// Mitsubishi GX Works2 project: Calculate   PLC: Q06UDEH (continued)

Import2Switch(ConveyorEntryIO:=Import2SwitchConveyorIn,
                          ConveyorExitIO:=Import2SwitchConveyorOut ,
                           SwitchIO:=Import2SwitchIO);
Import2SwitchIO.xLiftCylinderExtendButton:=M155;
Import2SwitchIO.xLiftCylinderRetractButton:=M156;
Y1ED:=Import2SwitchIO.xLiftCylinderExtend;
Y1EE:=Import2SwitchIO.xLiftCylinderRetract;
Import2SwitchIO.xLiftCylinderExtendDetect:=XF1;
Import2SwitchIO.xLiftCylinderRetractDetect:=XF2;
Import2SwitchConveyorIn.xCWPresent:=X104;
Import2SwitchConveyorIn.tLoadDelay:=T#2s;
Import2SwitchConveyorOut.xForward:=M149;
Import2SwitchConveyorOut.tLeaveDelay:=t#8s;
Import2SwitchConveyorOut.xCWPresent:=XF0;
Y1FC:=Import2SwitchConveyorIn.xMotorCW;

Import2LoadCylinder(ShuttleCarInOut:=Import2LoadCylinderIO);
ShuttleCarCurrentPosition( XF6 OR XF7 ,XF6 ,XF7, FALSE, Import2LoadCylinderIO.iCurrentPos );
Import2LoadCylinderIO.xReady:=TRUE;
Import2LoadCylinderIO.xForward:=M161;
Import2LoadCylinderIO.xBackward:=M162;
Import2LoadCylinderIO.xPosLimit:=TRUE;
Import2LoadCylinderIO.xNegLimit:=TRUE;
Y1ED:=Import2LoadCylinderIO.xCW;
Y1EE:=Import2LoadCylinderIO.xCCW;

(*2巷道出库*)
Export2Conveyor1(ConveyorMotor:=Export2Conveyor1IO);
Export2Conveyor1IO.tLeaveDelay:=t#10s;
Export2Conveyor1IO.xForward:=M96;
Export2Conveyor1IO.xCWPresent:=XFB;
Y1FD:=Export2Conveyor1IO.xMotorCW;

Export2Conveyor2(ConveyorMotor:=Export2Conveyor2iO);
Export2Conveyor2IO.tLeaveDelay:=t#10s;
Export2Conveyor2IO.xForward:=M97;
Export2Conveyor2IO.xCWPresent:=XFC;
Y1FE:=Export2Conveyor2IO.xMotorCW;

Export2Switch(ConveyorEntryIO:=Export2SwitchConveyorIn,
                          ConveyorExitIO:=Export2SwitchConveyorOut ,
                           SwitchIO:=Export2SwitchIO);
Export2SwitchIO.xLiftCylinderExtendButton:=M120;
Export2SwitchIO.xLiftCylinderRetractButton:=M121;
Export2SwitchIO.xLiftCylinderExtendInit:=1;
Y1F1:=Export2SwitchIO.xLiftCylinderExtend;
Y1F0:=Export2SwitchIO.xLiftCylinderRetract;
Export2SwitchIO.xLiftCylinderExtendDetect:=XF9;
Export2SwitchIO.xLiftCylinderRetractDetect:=XFA;
Export2SwitchConveyorIn.xForward:=M123;
Export2SwitchConveyorIn.xCWPresent:=X105;
Y1FF:=Export2SwitchConveyorIn.xMotorCW;
Export2SwitchConveyorOut.xCWPresent:=X105;

Export2LoadCylinder(ShuttleCarInOut:=Export2LoadCylinderIO);
ShuttleCarCurrentPosition( XFF OR XFE ,XFF ,XFE, FALSE, Export2LoadCylinderIO.iCurrentPos );
Export2LoadCylinderIO.xReady:=TRUE;
Export2LoadCylinderIO.xForward:=M124;
Export2LoadCylinderIO.xBackward:=M125;
Export2LoadCylinderIO.xPosLimit:=TRUE;
Export2LoadCylinderIO.xNegLimit:=TRUE;
Y1F2:=Export2LoadCylinderIO.xCW;
Y1F3:=Export2LoadCylinderIO.xCCW;

IF g_xAuto THEN
	(**高温库前自动程序**)
	Y187:=1;(***出库倍速链***)
(*	Y186:=1;(***入库倍速链***)
	IF  M883 AND XED THEN
        Export1LoadCylinderIO.xMDIExe:=1;
        Export1LoadCylinderIO.iDestinationPos:=1;
	END_IF;
	IF NOT XED THEN
        Export1LoadCylinderIO.xMDIExe:=1;
        Export1LoadCylinderIO.iDestinationPos:=2;
     END_IF;		
	Export1Conveyor1IO.xLoad:=XED AND Export1LoadCylinderIO.iCurrentPos=2;
	Export1Conveyor1IO.xUnload:=Export1Conveyor2IO.xEmpty;
	Export1Conveyor2IO.xLoad:=Export1Conveyor1IO.xNextRun;
	IF Y1E5 THEN
		Export1SwitchIO.xLiftCylinderExtendInit:=0;
	ELSE
		Export1SwitchIO.xLiftCylinderExtendInit:=1;
	END_IF;
	Export1Conveyor2Io.xUnload:=Export1SwitchConveyorIn.xEmpty;
	Export1SwitchIO.xEntryEnable:=Export1Conveyor2Io.xNextRun;
	Export1SwitchIO.xSwithEnable:=1;
	IF  M884 THEN
        Export2LoadCylinderIO.xMDIExe:=1;
        Export2LoadCylinderIO.iDestinationPos:=2;
	END_IF;
	Export2Conveyor1IO.xLoad:=XFD AND Export2LoadCylinderIO.iCurrentPos=2;
	Export2Conveyor1IO.xUnload:=Export2Conveyor2IO.xEmpty;
	Export2Conveyor2IO.xLoad:=Export2Conveyor1IO.xNextRun;
	Export2Conveyor2Io.xUnload:=Export2SwitchConveyorIn.xEmpty;
	Export2SwitchIO.xEntryEnable:=Export2Conveyor2Io.xNextRun;
	Export2SwitchIO.xSwithEnable:=1;
	
	H3000SwitchQuadPackageIO.xEntryEnable:=1;
	H3000SwitchQuadPackageIO.xSwithEnable:=1;
	H3000SwitchQuadPackageio.xExitEnable:=H3000Conveyor1IO.xEmpty;
	H3000Conveyor1Io.xLoad:=H3000SwitchPackageConveyorOut.xNextRun;
	H3000Conveyor1IO.xUnload:=H3000Conveyor2IO.xEmpty;
	H3000Conveyor2IO.xLoad:=H3000Conveyor1IO.xNextRun;
	H3000Conveyor2IO.xUnload:=H3000Conveyor3IO.xEmpty;
	H3000Conveyor3IO.xLoad:=H3000Conveyor2IO.xNextRun;	
	H3000Conveyor3IO.xUnload:=H3000Conveyor4IO.xEmpty;
	H3000Conveyor4IO.xLoad:=H3000Conveyor3IO.xNextRun;
	H3000Conveyor4IO.xUnload:=H3000Conveyor5IO.xEmpty;
	H3000Conveyor5IO.xLoad:=H3000Conveyor4IO.xNextRun;
	H3000Conveyor5IO.xUnload:=H3000Conveyor6IO.xEmpty;
	H3000Conveyor6IO.xLoad:=H3000Conveyor5IO.xNextRun;
	H3000Conveyor6IO.xUnload:=H3000Conveyor7IO.xEmpty;
	H3000Conveyor7IO.xLoad:=H3000Conveyor6IO.xNextRun;
	H3000Conveyor7IO.xUnload:=H3000Conveyor8IO.xEmpty;
	H3000Conveyor8IO.xLoad:=H3000Conveyor7IO.xNextRun;	
	H3000Conveyor8IO.xUnload:=H3000Conveyor9IO.xEmpty;
	H3000Conveyor9IO.xLoad:=H3000Conveyor8IO.xNextRun;	
	H3000Conveyor9IO.xUnload:=H3000Conveyor10IO.xEmpty;
	H3000Conveyor10IO.xLoad:=H3000Conveyor9IO.xNextRun;
	H3000Conveyor10IO.xUnload:=D401.0;
	D201.0:=H3000Conveyor10IO.xNextRun;

	
	(*H2200Conveyor1IO.xLoad:=;*)
	H2200Conveyor1IO.xUnload:=H2200Conveyor2IO.xEmpty;
	H2200Conveyor2IO.xLoad:=H2200Conveyor1IO.xNextRun;
	H2200Conveyor2IO.xUnload:=H2200Conveyor3IO.xEmpty;
	H2200Conveyor3IO.xLoad:=H2200Conveyor2IO.xNextRun;	
	H2200Conveyor3IO.xUnload:=H2200Conveyor4IO.xEmpty;
	H2200Conveyor4IO.xLoad:=H2200Conveyor3IO.xNextRun;
	H2200Conveyor4IO.xUnload:=H2200Conveyor5IO.xEmpty;
	H2200Conveyor5IO.xLoad:=H2200Conveyor4IO.xNextRun;
	H2200Conveyor5IO.xUnload:=H2200Conveyor6IO.xEmpty;
	H2200Conveyor6IO.xLoad:=H2200Conveyor5IO.xNextRun;
	H2200Conveyor6IO.xUnload:=H2200Conveyor7IO.xEmpty;
	H2200Conveyor7IO.xLoad:=H2200Conveyor6IO.xNextRun;
	H2200Conveyor7IO.xUnload:=H2200Conveyor8IO.xEmpty;
	H2200Conveyor8IO.xLoad:=H2200Conveyor7IO.xNextRun;	
	H2200Conveyor8IO.xUnload:=H2200Conveyor9IO.xEmpty;
	H2200Conveyor9IO.xLoad:=H2200Conveyor8IO.xNextRun;	
	H2200Conveyor9IO.xUnload:=H2200Conveyor10IO.xEmpty;
	H2200Conveyor10IO.xLoad:=H2200Conveyor9IO.xNextRun;
	H2200Conveyor10IO.xUnload:=D401.1;
	D201.1:=H2200Conveyor10IO.xNextRun;
	(*化成回流线体*)
	D201.2:=H1000Conveyor10IO.xEmpty;
	H1000Conveyor10IO.xLoad:=D401.2;
	H1000Conveyor10IO.xUnload:=H1000Conveyor9IO.xEmpty;
    H1000Conveyor9IO.xLoad:=H1000Conveyor10IO.xNextRun;
    H1000Conveyor9IO.xUnload:=H1000Conveyor8IO.xEmpty;
    H1000Conveyor8IO.xLoad:=H1000Conveyor9IO.xNextRun;
    H1000Conveyor8IO.xUnload:=H1000Conveyor7IO.xEmpty;
    H1000Conveyor7IO.xLoad:=H1000Conveyor8IO.xNextRun;
    H1000Conveyor7IO.xUnload:=H1000Conveyor6IO.xEmpty;
    H1000Conveyor6IO.xLoad:=H1000Conveyor7IO.xNextRun;
    H1000Conveyor6IO.xUnload:=H1000Conveyor5IO.xEmpty;
    H1000Conveyor5IO.xLoad:=H1000Conveyor6IO.xNextRun;
    H1000Conveyor5IO.xUnload:=H1000Conveyor4IO.xEmpty;
    H1000Conveyor4IO.xLoad:=H1000Conveyor5IO.xNextRun;
    H1000Conveyor4IO.xUnload:=H1000Conveyor3IO.xEmpty;
    H1000Conveyor3IO.xLoad:=H1000Conveyor4IO.xNextRun;
    H1000Conveyor3IO.xUnload:=H1000Conveyor2IO.xEmpty;
    H1000Conveyor2IO.xLoad:=H1000Conveyor3IO.xNextRun;  
    H1000Conveyor2IO.xUnload:=H1000Conveyor1IO.xEmpty;
    H1000Conveyor1IO.xLoad:=H1000Conveyor2IO.xNextRun; 
    IF H1000Conveyor1IO.xEmpty=0 AND Lifter2Occupy=0 THEN
    	Lifter2IO.xMDIExe:=1;
    	Lifter2IO.iDestinationPos:=2;
    END_IF;    
    IF Lifter2IO.iCurrentPos=2 AND (D190-Lifter2Position[Lifter2IO.iDestinationPos])<10  THEN 
    	H1000Conveyor1IO.xUnload:=Conveyor2IO.xEmpty;
    	Conveyor2IO.xloadCCW:=1;
    ELSE
    	H1000Conveyor1IO.xUnload:=0;
    END_IF;
    	Conveyor2IO.xLoad:=H1000Conveyor1IO.xNextRun;     
	(*注液设备满框入库*)
	H850Conveyor4IO.xLoad:=M880;
	H850Conveyor4IO.xUnload:=H850Conveyor5IO.xEmpty;
	H850Conveyor5IO.xLoad:=H850Conveyor4IO.xNextRun;
	H850Conveyor5IO.xUnload:=H850Conveyor6IO.xEmpty;
	H850Conveyor6IO.xLoad:=H850Conveyor5IO.xNextRun;	
	IF H850RotorConveyorIO.xEmpty THEN
		 H850RotorIO.xMDIExe:=1;
		  H850RotorIO.iDestinationPos:=1;
	END_IF;
	IF H850RotorConveyorIO.xEmpty=0 THEN
		 H850RotorIO.xMDIExe:=1;
		  H850RotorIO.iDestinationPos:=2;
	END_IF;	
	IF H850RotorIO.iCurrentPos=1 THEN
    H850Conveyor6IO.xUnload:=H850RotorConveyorIO.xEmpty;
	ELSE
	 H850Conveyor6IO.xUnload:=0;
	END_IF;	
	H850RotorConveyorIO.xLoad:=H850Conveyor6IO.xNextRun;
	IF H850RotorIO.iCurrentPos=2 THEN
		H850RotorConveyorIO.xUnload:=H850SwitchConveyorIn.xEmpty AND H850SwitchConveyorOut.xEmpty;
	ELSE
		H850RotorConveyorIO.xUnload:=0;
	END_IF;
	H850SwitchIO.xEntryEnable:=H850RotorConveyorIO.xNextRun;	
	H850SwitchIO.xSwithEnable:=1;
	H850SwitchIO.xExitEnable:=H850Conveyor8IO.xEmpty;
    H850Conveyor8IO.xLoad:=H850SwitchConveyorOut.xNextRun;
    
    IF H850Conveyor8IO.xEmpty=0 AND NOT Lifter2Occupy THEN
    	Lifter2IO.xMDIExe:=1;
    	Lifter2IO.iDestinationPos:=1;
    END_IF;
    IF Lifter2IO.iCurrentPos=1 AND ABS(D190-Lifter2Position[Lifter2IO.iDestinationPos])<10 THEN
    	H850Conveyor8IO.xUnload:= Conveyor2IO.xEmpty;
    	Conveyor2IO.xLoad:=H850Conveyor8IO.xNextRun;
        Conveyor2IO.xloadCCW:=0;
    ELSE
    	H850Conveyor8IO.xUnload:=0;
    END_IF;
     IF NOT Lifter2ExportChem AND Conveyor2IO.xEmpty=0 THEN(*只要不是加压化成的 满框都要入库*)
     	Lifter2IO.xMDIExe:=1;
    	Lifter2IO.iDestinationPos:=3;
     END_IF;
    IF Lifter2IO.iCurrentPos=3 AND ABS(D190-Lifter2Position[Lifter2IO.iDestinationPos])<10 THEN	
		Conveyor2IO.xUnload:=H2200ImportConveyor2IO.xEmpty;
		H2200ImportConveyor2IO.xLoad:=Conveyor2IO.xNextRun;  
		Conveyor2IO.xUnloadCCW:=1;  	
    END_IF;
    (*不在目标位置不可下料*)
    IF ABS(D190-Lifter2Position[Lifter2IO.iDestinationPos])>10 THEN
    	Conveyor2IO.xUnload:=0;
    END_IF;
    H2200ImportConveyor2IO.xUnload:=H2200Switch1ConveyorOut.xEmpty;
    H2200Switch1ConveyorOut.xLoad:=H2200ImportConveyor2IO.xNextRun;
    IF LDP(TRUE,  NOT H2200ImportConveyor2IO.xEmpty ) THEN
    H2200Switch1IO.xLiftCylinderExtendInit:=1;
    END_IF;
    H2200ImportConveyor1IO.xLoad:=H2200Switch1ConveyorOut.xNextRun;
    H2200Switch1ConveyorOut.xUnload:=H2200ImportConveyor1IO.xEmpty;
    
    H2200ImportConveyor1IO.xUnload:=H2200Switch2ConveyorIn.xEmpty;
    H2200Switch2IO.xEntryEnable:=H2200ImportConveyor1IO.xNextRun;
    H2200Switch2IO.xSwithEnable:=1;
    H2200Switch2IO.xExitEnable:=1;
    
    Import1SwitchIO.xEntryEnable:=1;
    Import1SwitchIO.xSwithEnable:=1;
    Import1SwitchIO.xExitEnable:=Import1Conveyor1IO.xEmpty;
    Import1Conveyor1IO.xLoad:=Import1SwitchConveyorOut.xNextRun;
    Import1Conveyor1IO.xUnload:=Import1Conveyor2IO.xEmpty AND NOT XE5;
    Import1Conveyor2IO.xLoad:=Import1Conveyor1IO.xNextRun;
    
    IF Import1Conveyor2IO.xEmpty=0 AND XE5 THEN
    	Import1LoadCylinderIO.xMDIExe:=1;
    	Import1LoadCylinderIO.iDestinationPos:=2;
    	Import1Conveyor2IO.xPutInto:=0;
    END_IF;
    IF NOT XE5 THEN
    	Import1LoadCylinderIO.xMDIExe:=1;
    	Import1LoadCylinderIO.iDestinationPos:=1;
    	Import1Conveyor2IO.xPutInto:=1;
    END_IF;
    
    Y173:=1;(*空框A返回倍速链*)
   Y175:=1;(*空框B返回倍速链*)
   (*空框回流*)
   H2200SwitchEmptyABackIO.xEntryEnable:=1;
   H2200SwitchEmptyABackIO.xLiftCylinderExtendInit:=1;
    H2200SwitchEmptyABackIO.xSwithEnable:=1;
    H2200SwitchEmptyABackIO.xExitEnable:=H2200RotorConveyorIO.xEmpty AND H2200RotorIO.iCurrentPos=1 AND X6F;
    IF ldp(TRUE,H2200SwitchEmptyABackConveyorIn.xEmpty=0) THEN
    	H2200Switch1IO.xLiftCylinderExtendInit:=0;
    END_IF;
    IF H2200RotorConveyorIO.xEmpty THEN
    	H2200RotorIO.xMDIExe:=1;
    	H2200RotorIO.iDestinationPos:=1;
    END_IF;
    IF H2200RotorConveyorIO.xEmpty=0 THEN
     	H2200RotorIO.xMDIExe:=1;
    	H2200RotorIO.iDestinationPos:=2;   
    END_IF;   
    IF H2200RotorIO.iCurrentPos=1 AND X6F THEN
    	H2200RotorConveyorIO.xLoad:=H2200SwitchEmptyABackConveyorOut.xNextRun OR H2200SwitchEmptyBBackConveyorOut.xNextRun;
    	H2200SwitchEmptyABackIO.xExitEnable:=H2200RotorConveyorIO.xEmpty;
    	H2200SwitchEmptyBBackIO.xExitEnable:=H2200RotorConveyorIO.xEmpty;
    ELSE
     	H2200SwitchEmptyABackIO.xExitEnable:=0;
    	H2200SwitchEmptyBBackIO.xExitEnable:=0;   
    	H2200RotorConveyorIO.xLoad:=0;	
    END_IF;
    IF Conveyor1IO.xEmpty THEN
    	Lifter1IO.xMDIExe:=1;
    	Lifter1IO.iDestinationPos:=2;
    END_IF;
    IF Conveyor1IO.xEmpty=0 THEN
    	Lifter1IO.xMDIExe:=1;
    	Lifter1IO.iDestinationPos:=1; 
    END_IF;
    IF Lifter1IO.iCurrentPos=2 AND X8D AND H2200RotorIO.iCurrentPos=2 AND X75 THEN
    	H2200RotorConveyorIO.xUnload:=Conveyor1IO.xEmpty;
    ELSE
    	H2200RotorConveyorIO.xUnload:=0;
    END_IF;
    Conveyor1IO.xLoad:=H2200RotorConveyorIO.xNextRun; 
    IF Lifter1IO.iCurrentPos=1 AND X8C THEN
    	Conveyor1IO.xUnload:=H850Conveyor3IO.xEmpty;
    ELSE
    	Conveyor1IO.xUnload:=0;
    END_IF;  	
    H850Conveyor3IO.xLoad:=Conveyor1IO.xNextRun;
    h850conveyor3IO.xUnload:=H850Conveyor1IO.xEmpty;
    H850Conveyor1IO.xLoad:=H850Conveyor3IO.xNextRun;
END_IF;

IF g_xManual THEN
    D201:=0;(*发送给化成B柜*)
	IF M134 THEN (*空框A返回倍速链 手动*)
		 Y173:=1;(*空框A返回倍速链*)
	ELSE
		Y173:=0;;(*空框A返回倍速链*)
	END_IF;
	IF M135 THEN (*空框B返回倍速链 手动*)
		 Y175:=1;(*空框B返回倍速链*)
	ELSE
		Y175:=0;(*空框B返回倍速链*)
	END_IF;	
	IF M163 THEN (*入库倍速链 手动*)
		 Y186:=1;(*入库倍速链*)
	ELSE
		Y186:=0;;(*入库倍速链*)
	END_IF;
	IF M64 THEN (*出库倍速链 手动*)
		 Y187:=1;(*出库倍速链 *)
	ELSE
		Y187:=0;(*出库倍速链 *)
	END_IF;		
END_IF;
END_PROGRAM

PROGRAM Start
IF g_xReset THEN
	SM50:=1;
ELSE
	SM50:=0;
END_IF;
CASE g_iState OF
	0: 
		g_xManual:=1;
		g_xAuto:=0;	
		g_xStackLampAmber:=1;
		g_xStackLampGreen:=0;
		g_xRemoteAuto:=0;
	1:
		g_xManual:=0;
		g_xAuto:=1;
		g_xStackLampGreen:=1;
		g_xStackLampAmber:=0;
		g_xRemoteAuto:=0;
	2:	
        g_xRemoteAuto:=1;
        g_xStackLampGreen:=1;
        g_xStackLampAmber:=0;
        g_xAuto:=0;
		g_xManual:=0;
END_CASE;
IF g_xLocalAutoStart THEN  
	g_iState:=1;
END_IF;

IF g_xStop OR g_xEStop=0 THEN 
	g_iState:=0;
END_IF;
IF g_xRemoteAutoStart THEN
	g_iState:=2;
END_IF;
END_PROGRAM

PROGRAM UDP
(*与化成柜2通讯*)
D200:=2;
SP_SOCOPEN( SM403 AND NOT SD1282.0 AND NOT SD1284.0 AND SD1288.A , "U0", K1 , D110 , M100);
SP_SOCSND( SM413 AND SD1282.0 , "U0" , K1 , D100, D200, M102 );
SP_SOCRCV( SD1282.0 AND SD1286.0 AND NOT M104 , "U0" , K1, D300 , D400 ,M104 );
SP_SOCCLOSE( LDF(TRUE,SD1082.0) , "U0" , K1, D120, M106 );
(*编码器处理程序*)
IF XA OR X0B   THEN
	D140:=2;
	D143:=6;
END_IF;
	G_INPUT( X0A OR X0B, 0 , D140 , D160 , M110 );(*串口数据读取指令*)
IF M110 THEN
	D170:=0;
	D172:=4;
END_IF;
ZP_CSET( M110  , "U0", 2 , D170, D180,M112 );(*串口数据缓存区清除指令*)
IF D160=11069 THEN  (*接收到数据开始执行ASCII码转换成10进制，D160为=+ ，串口传输的字头 转换为10进制是11069，不判断这个报4100错误*)
    DABIN( TRUE , D163, D190 );
END_IF;
END_PROGRAM

FUNCTION_BLOCK Conveyor
VAR
  tRundelay : TIME;  (* 离开延时 *)
END_VAR
VAR_IN_OUT
  ConveyorMotor : ConveyorIO;  (* 输送线输入输出 *)
END_VAR
VAR
  iStep : INT;  (* 上料步骤 *)
  m_tLoadTimer : TIME;  (* 上料计时器 *)
  m_tUnloadTimer : TIME;  (* 下料计时器 *)
  m_tonLeaveDelay : TON;  (* 离开延时定时器 *)
  m_xLeaveDelayOut : BOOL;  (* 离开延时 *)
  m_tLeaveCurrentTime : TIME;
  m_tonLoadAlarm : TON;  (* 上料延时报警 *)
END_VAR
VAR CONSTANT
  LOAD_UNLOAD_TIME : TIME := T#30s;  (* 延时报警常量 *)
END_VAR
VAR
  m_tonUnloadAlam : TON;  (* 下料报警定时器 *)
  m_tonLoadDelay : TON;  (* 上料延时 *)
  m_xLoadDelayOut : BOOL;  (* 上料延时输出 *)
  m_tLoadCurrentTime : TIME;  (* 上料延时当前时间 *)
  m_xInitial : BOOL;  (* 初始化 *)
END_VAR
(*////////////////////////////////////////////////////////////////////////////////////////////////////////////
//传输线控制FB块，可控制单方向线体，双向旋转线体，支持双向上下料            
//线体初始化后为空的情况下输入xLoad信号即可进行上料动作，使用xLoadCCW信号可反方向上料
//增加了产品信息和产品种类的储存，当传输线为空和上料进行标志位为零的情况下清除产品信息和产品种类
//使用方式是在置位xLoad信号后，把产品信息和产品种类传入，等下料后自动清零
//线体不为空的情况下使用xUnload信号可进行下料动作，物料有无传感器的下降沿后出发计时器，延时断开传输线旋转
//单方向传输线体把xLoadCCW、xUnloadCCW设置为零，双向线体上料方向和下料反向的,方向固定的 把xUnloadCCW设置为1
//双方向线体双向都能上下料的要根据上料的方向来设置xLoadCCW,xUnloadCCW
//增加工作中信号xBusy当电机正转 显示为工作中
//增加上下料超时报警，xLoadAlarm，xUnloadAlarm，设定时间在LOAD_UNLOAD_TIME常量上，现在设置的为30秒
//增加xPutInto信号，用于直接投入的物料，检测开关感应到后，直接进入下料流程，上升沿有效
//离开延时改为变量 iLeaveDelay 默认为0 离开检测开关离输送线尾端比较远的线体需要根据情况设定100ms为单位
增加初始化标志位，增加进入延时时间，初始化为进入延时时间为0 ，离开延时时间为2S，通过外围接口可以更改
//修改信息  修改后请增加版本
//YAO      V1.0
///////////////////////////////////////////////////////////////////////////////////////////////////////////
********************************************************)
IF NOT m_xInitial THEN
	ConveyorMotor.tLoadDelay:=T#0s;
	ConveyorMotor.tLeaveDelay:=T#2s;
END_IF;
m_xInitial:=1;
IF g_xAuto THEN
CASE iStep OF
	0:
	ConveyorMotor.xMotorCW:=0;
	ConveyorMotor.xMotorCCW:=0;
	ConveyorMotor.xNextRun:=0;
IF g_xEStop  THEN
	IF (ConveyorMotor.xCWPresent OR ConveyorMotor.xCCWPresent)  THEN
		iStep:=3;
		ConveyorMotor.xEmpty:=0;
		ELSE
		iStep:=1;
		ConveyorMotor.xEmpty:=1;
	END_IF;
END_IF;		
	1: 
	IF ConveyorMotor.xLoad    
		AND ConveyorMotor.xMotorCW=0   
		AND ConveyorMotor.xMotorCCW=0   
		AND ConveyorMotor.xEmpty THEN	
		iStep:=2;
	END_IF;
	2: 
	IF ConveyorMotor.xloadCCW THEN
		ConveyorMotor.xMotorCCW:=1; 
		ConveyorMotor.xMotorCW:=0;
	ELSE
	    ConveyorMotor.xMotorCW:=1;  
		ConveyorMotor.xMotorCCW:=0;
	END_IF;
		m_tonLoadDelay(IN:= (ConveyorMotor.xCWPresent AND NOT ConveyorMotor.xloadCCW) 
		                                        OR (ConveyorMotor.xCCWPresent AND ConveyorMotor.xloadCCW) ,
		                               PT:= ConveyorMotor.tLoadDelay ,
		                               Q:= m_xLoadDelayOut ,
		                               ET:= m_tLoadTimer );
	    IF m_xLoadDelayOut THEN 	 
		    iStep:=3;
		END_IF;
	3:
	ConveyorMotor.xMotorCW:=0;
	ConveyorMotor.xMotorCCW:=0;
	ConveyorMotor.xEmpty:=0;
	IF ConveyorMotor.xUnload THEN 
		iStep:=4;
	END_IF;
	4:	
	IF ConveyorMotor.xUnloadCCW THEN   
		ConveyorMotor.xMotorCCW:=1;  
		ConveyorMotor.xMotorCW:=0;

		ConveyorMotor.xLeave:=ldf(TRUE,ConveyorMotor.xCCWPresent) OR ConveyorMotor.xLeave;
		ELSE
	    ConveyorMotor.xMotorCW:=1;  
		ConveyorMotor.xMotorCCW:=0;
		ConveyorMotor.xLeave:=ldf(TRUE,ConveyorMotor.xCWPresent) OR ConveyorMotor.xLeave;
	END_IF;
	ConveyorMotor.xNextRun:=1; 
	m_tonLeaveDelay(IN:= ConveyorMotor.xLeave,PT:= ConveyorMotor.tLeaveDelay,Q:=m_xLeaveDelayOut ,ET:= m_tLeaveCurrentTime );	
	IF m_xLeaveDelayOut THEN
		ConveyorMotor.xMotorCW:=0;
		ConveyorMotor.xMotorCCW:=0;
		iStep:=0;
		ConveyorMotor.xNextRun:=0;
		ConveyorMotor.xLeave:=0;
		ConveyorMotor.xEmpty:=1;		
	END_IF;	
	IF NOT ConveyorMotor.xUnload THEN 
		istep:=0;
	END_IF;
END_CASE;
IF LDP(TRUE,ConveyorMotor.xPutInto) THEN
	iStep:=0;
END_IF;
END_IF;
IF ConveyorMotor.xEmpty AND NOT ConveyorMotor.xLoad THEN
	ConveyorMotor.iProductCategory:=0;
END_IF;
IF g_xEStop=0 OR g_xReset THEN
	iStep:=0;
END_IF;	

IF g_xManual THEN
	iStep:=0;

	IF ConveyorMotor.xForward 
		AND ConveyorMotor.xBackward=0 
		AND ConveyorMotor.xMotorCCW=0
		AND g_xEStop THEN
		ConveyorMotor.xMotorCW:=1;
		ConveyorMotor.xMotorCCW:=0;
		ELSE
		ConveyorMotor.xMotorCW:=0;
	END_IF;

	IF ConveyorMotor.xBackward 
		AND ConveyorMotor.xForward=0 
		AND ConveyorMotor.xMotorCW=0
		AND g_xEStop  THEN
		ConveyorMotor.xMotorCCW:=1;
		conveyormotor.xMotorCW:=0;
		ELSE
		ConveyorMotor.xMotorCCW:=0;
	END_IF;
END_IF;
IF ConveyorMotor.xMotorCCW        
	OR ConveyorMotor.xMotorCW THEN  
	ConveyorMotor.xBusy:=1;
	ELSE
	ConveyorMotor.xBusy:=0;
END_IF;
m_tonLoadAlarm(IN:= iStep=2 ,PT:= LOAD_UNLOAD_TIME,Q:= ConveyorMotor.xLoadAlarrm ,ET:= m_tLoadTimer );
m_tonUnloadAlam(IN:= iStep=4,PT:= LOAD_UNLOAD_TIME,Q:= ConveyorMotor.xUnloadAlarm,ET:= m_tUnloadTimer );
END_FUNCTION_BLOCK

FUNCTION_BLOCK ShuttleCar
VAR_IN_OUT
  ShuttleCarInOut : ShuttleCarIO;
END_VAR
VAR
  m_xBrakeDelay : BOOL;  (* 刹车延时标志位 *)
  diCurrentPosRetain : DINT;
  m_tonBrakeDelay : TON;  (* 延时 *)
  m_tBrakeDelay : TIME;
  m_xBrake : BOOL;
  m_tBrakeDelayCurrentTime : TIME;
END_VAR
(*******************************************************************
输送小车程序，可用于使用认址片控制位置的输送车程序，可用于控制提升机，
使用了限位捕捉程序防止小车惯性过大冲过限位后继续行走，捕捉程序采用反
转复位，这样设计有弊端可能反转复位后车的位置并没有回到限位以内,当两个
限位同时碰到的时候，会使运料小车进入死锁状态，通过xPassLimit来解开死锁，
可以在触摸屏中使用一个带权限的按钮来进行控制，配合ShuttleCarCurrentPos
函数来计算位置信息
修改信息  修改后请增加版本
YAO      V1.0
********************************************************************)

ShuttleCarInOut.xPosLimitCatch:=LDF(TRUE,ShuttleCarInOut.xPosLimit) OR ShuttleCarInOut.xPosLimitCatch;
IF ShuttleCarInOut.xCCW THEN  
	ShuttleCarInOut.xPosLimitCatch:=0;
END_IF;

ShuttleCarInOut.xNegLimitCatch:=LDF(TRUE,ShuttleCarInOut.xNegLimit) OR ShuttleCarInOut.xNegLimitCatch;
IF ShuttleCarInOut.xCW THEN   
	ShuttleCarInOut.xNegLimitCatch:=0;  
END_IF;
IF ShuttleCarInOut.xPassLimit OR
	(ShuttleCarInOut.xNegLimitCatch 
	AND ShuttleCarInOut.xPosLimitCatch)  THEN  
	ShuttleCarInOut.xNegLimitCatch:=0; 
	ShuttleCarInOut.xPosLimitCatch:=0;
END_IF;

IF ShuttleCarInOut.xReady THEN	
    IF g_xManual THEN  
	    IF ShuttleCarInOut.xForward 
			AND ShuttleCarInOut.xBackward=0 
			AND ShuttleCarInOut.xCCW=0 
			AND ShuttleCarInOut.xPosLimitCatch=0 
			AND g_xEStop THEN
		    ShuttleCarInOut.xCW:=1;
		    ELSE
		    ShuttleCarInOut.xCW:=0;
	    END_IF;
	    IF ShuttleCarInOut.xBackward 
			AND ShuttleCarInOut.xForward=0 
			AND ShuttleCarInOut.xCW=0 
			AND ShuttleCarInOut.xNegLimitCatch=0 
			AND G_xEStop THEN  
		    ShuttleCarInOut.xCCW:=1;
		    ELSE
		    ShuttleCarInOut.xCCW:=0;
	    END_IF;
    END_IF;
  IF g_xAuto AND g_xEStop THEN  
	  IF ShuttleCarInOut.xMDIExe AND ShuttleCarInOut.iDestinationPos<>0 THEN
	
	    IF ShuttleCarInOut.iCurrentPos<ShuttleCarInOut.iDestinationPos AND ShuttleCarInOut.xPosLimitCatch=0 THEN
			ShuttleCarInOut.xCW:=1;
			ShuttleCarInOut.xCCW:=0;
			ShuttleCarInOut.xMDIDone:=0;
		END_IF;

		IF ShuttleCarInOut.iCurrentPos>ShuttleCarInOut.iDestinationPos AND ShuttleCarInOut.xNegLimitCatch=0 THEN
			ShuttleCarInOut.xCCW:=1;
			ShuttleCarInOut.xCW:=0;
			ShuttleCarInOut.xMDIDone:=0;
		END_IF;
	
		IF ShuttleCarInOut.iCurrentPos=ShuttleCarInOut.iDestinationPos THEN
			ShuttleCarInOut.xCW:=0;
			ShuttleCarInOut.xCCW:=0;
			ShuttleCarInOut.xMDIDone:=1;
			ELSE
			ShuttleCarInOut.xMDIDone:=0;
		END_IF;

		IF ShuttleCarInOut.xPosLimitCatch THEN
			ShuttleCarInOut.xCW:=0;
			ShuttleCarInOut.xMDIDone:=0;
		END_IF;

		IF ShuttleCarInOut.xNegLimitCatch THEN
			ShuttleCarInOut.xCCW:=0;
			ShuttleCarInOut.xMDIDone:=0;
		END_IF;
		ELSE
		ShuttleCarInOut.xCW:=0;
		ShuttleCarInOut.xCCW:=0;
		ShuttleCarInOut.xMDIDone:=0;
	  END_IF;
	END_IF;
	ELSE
		ShuttleCarInOut.xCW:=0;
		ShuttleCarInOut.xCCW:=0;	
END_IF;

m_tonBrakeDelay(IN:=m_xBrakeDelay ,PT:= T#100ms,Q:=m_xBrake ,ET:= m_tBrakeDelayCurrentTime);
IF (ShuttleCarInOut.xCW OR ShuttleCarInOut.xCCW) AND ShuttleCarInOut.xReady=1 THEN
	ShuttleCarInOut.xBrake:=m_xBrake;
	m_xBrakeDelay:=1;
	ELSE
	ShuttleCarInOut.xBrake:=0;
	m_xBrakeDelay:=0;
END_IF;

IF g_xEStop =0 THEN
	ShuttleCarInOut.xCW :=0;
	ShuttleCarInOut.xCCW:=0;
END_IF;

(*IF SM402 THEN 
	ShuttleCarInOut.diCurrentPos:=diCurrentPosRetain;
	ELSE
	diCurrentPosRetain:=ShuttleCarInOut.diCurrentPos;
END_IF;*)

IF ShuttleCarInOut.xCW OR ShuttleCarInOut.xCCW THEN
	ShuttleCarInOut.xBusy:=1;
	ELSE
	ShuttleCarInout.xBusy:=0;
END_IF;
END_FUNCTION_BLOCK

FUNCTION ShuttleCarCurrentPosition
VAR_INPUT
  xPosition1 : BOOL;
  xPosition2 : BOOL;
  xPosition3 : BOOL;
END_VAR
(************************************
计算输送车当前位置的函数
**************************************)
IF xPosition1 THEN
	ShuttleCarCurrentPosition:=1;
END_IF;
IF xPosition2 THEN
	ShuttleCarCurrentPosition:=2;
END_IF;
IF xPosition3 THEN
	ShuttleCarCurrentPosition:=3;
END_IF;
END_FUNCTION

FUNCTION_BLOCK Switch
VAR_IN_OUT
  ConveyorEntryIO : ConveyorIO;
END_VAR
VAR
  ConveyorEntry : Conveyor;
  m_tonEntryBarDelay : TON;  (* 进入阻挡器延时 *)
  m_tEntryBarDelay : TIME;
  m_xEntryBarDelay : BOOL;
END_VAR
VAR_IN_OUT
  ConveyorExitIO : ConveyorIO;
END_VAR
VAR
  m_tonLiftCylinderDelay : TON;  (* 顶升延时 *)
  m_xLiftCylinderDelay : BOOL;
  m_tLiftCylinderDelay : TIME;
  m_tonExitBarDelay : TON;  (* 退出阻挡器延时 *)
  m_tExitBarDelay : TIME;
  m_xExitBarDelay : BOOL;
END_VAR
VAR_IN_OUT
  SwitchIO : SwitchIO;
END_VAR
VAR
  iStep : INT;
  ConveyorExit : Conveyor;
  m_xInitial : BOOL;
END_VAR
ConveyorEntry(ConveyorMotor:=ConveyorEntryIO);
ConveyorExit(ConveyorMotor:=ConveyorExitIO);

IF NOT m_xInitial THEN
	ConveyorExitIO.tLeaveDelay:=T#5s;
END_IF;
m_xInitial:=1;

IF g_xAuto THEN
	CASE iStep OF
		0:(*初始化*)
		ConveyorEntryIO.xLoad:=0;
		ConveyorEntryIO.xUnload:=0;
		ConveyorEntryIO.xPutInto:=0;
		ConveyorExitIO.xLoad:=0;
		ConveyorExitIo.xUnload:=0;
		ConveyorExitIO.xPutInto:=0;
		SwitchIO.xEntryBarCylinderRetract:=0;
		SwitchIO.xExitBarCylinderRetract:=0;
		IF SwitchIO.xLiftCylinderExtendInit THEN
			SwitchIO.xLiftCylinderExtend:=1;
			SwitchIO.xLiftCylinderRetract:=0;
		    IF SwitchIO.xLiftCylinderExtendDetect THEN
			    iStep:=1;
		     END_IF; 
		ELSE
			SwitchIO.xLiftCylinderExtend:=0;
			SwitchIO.xLiftCylinderRetract:=1;	
		    IF SwitchIO.xLiftCylinderRetractDetect THEN
			    iStep:=1;
		    END_IF;		
		END_IF;
		1:(*上料*)
        IF SwitchIO.xEntryEnable AND ConveyorEntryIO.xEmpty AND ConveyorExitIO.xEmpty THEN
        	SwitchIO.xEntryBarCylinderRetract:=1;
        	ConveyorEntryIO.xLoad:=1;
        END_IF;
        m_tonEntryBarDelay(IN:=SwitchIO.xEntryBarCylinderRetract ,PT:=T#1S ,Q:= m_xEntryBarDelay ,ET:= m_tEntryBarDelay );
        IF m_xEntryBarDelay THEN
        	ConveyorEntryIO.xPutInto:=1;
        END_IF;
        IF ConveyorEntryIO.xEmpty=0 THEN
        	SwitchIO.xEntryBarCylinderRetract:=0;
        	ConveyorEntryIO.xLoad:=0;
        	ConveyorExitIO.xPutInto:=1;
        END_IF;
        IF m_xLiftCylinderDelay AND  SwitchIO.xSwithEnable THEN
        	 iStep:=2;
        END_IF;
        IF SwitchIO.xSwithEnable=0 AND m_xLiftCylinderDelay  THEN
        	 iStep:=3;
        END_IF;
		2:(*顶升*)
			SwitchIO.xExitBarCylinderRetract:=0;
			ConveyorEntryIO.xPutInto:=0;(*复位进入初始化*)
		    IF SwitchIO.xLiftCylinderExtendInit THEN
			    SwitchIO.xLiftCylinderExtend:=0;
			    SwitchIO.xLiftCylinderRetract:=1;
		    ELSE
			    SwitchIO.xLiftCylinderExtend:=1;
			    SwitchIO.xLiftCylinderRetract:=0;			
		   END_IF;

		  IF SwitchIO.xLiftCylinderExtendInit THEN
		  	IF SwitchIO.xLiftCylinderRetractDetect THEN
		  		iStep:=4;
		  	END_IF;
		  	ELSE
		  	IF SwitchIO.xLiftCylinderExtendDetect THEN
		      iStep:=4; 
		  	END_IF;
		  END_IF;
		  3:(*放行*)	
		  	SwitchIO.xExitBarCylinderRetract:=1;
		  	iStep:=4;
		  4:(*下料*)
		  IF SwitchIO.xExitEnable  AND m_xExitBarDelay THEN		  
		  ConveyorExitIO.xUnload:=1;
		  END_IF;
		  IF ConveyorExitIO.xEmpty OR ConveyorEntryIO.xEmpty  THEN
		  	COnveyorExitIO.xUnload:=0;
		  	ConveyorExitIO.xPutInto:=1;
		  	ConveyorEntryIO.xPutInto:=1;
			iStep:=0; 
		  END_IF;
	END_CASE;
        m_tonLiftCylinderDelay(IN:=NOT ConveyorEntryIO.xEmpty AND iStep=1 ,PT:= T#1S ,Q:= m_xLiftCylinderDelay ,ET:=m_tLiftCylinderDelay );
 		m_tonExitBarDelay(IN:=iStep=4 ,PT:= T#1s ,Q:= m_xExitBarDelay ,ET:= m_tExitBarDelay);
END_IF;
IF g_xReset OR LDP(TRUE,SwitchIO.xLiftCylinderExtendInit) OR LDF(TRUE,SwitchIO.xLiftCylinderExtendInit) THEN
	iStep:=0;
END_IF;
IF g_xManual  THEN
	iStep:=0;
	ConveyorEntryIO.xLoad:=0;
    ConveyorEntryIO.xUnload:=0;
	ConveyorEntryIO.xPutInto:=0;
	ConveyorExitIO.xLoad:=0;
	ConveyorExitIo.xUnload:=0;
	ConveyorExitIO.xPutInto:=0;
	SwitchIO.xEntryBarCylinderRetract:=0;
	SwitchIO.xExitBarCylinderRetract:=0;
	IF SwitchIO.xEntryBarCylinderRetractButton THEN
		SwitchIO.xEntryBarCylinderRetract:=1;
	ELSE
		SwitchIO.xEntryBarCylinderRetract:=0;
	END_IF;
		IF SwitchIO.xExitBarCylinderRetractButton THEN
		SwitchIO.xExitBarCylinderRetract:=1;
	ELSE
		SwitchIO.xExitBarCylinderRetract:=0;
		END_IF;
		IF SwitchIO.xLiftCylinderExtendButton AND NOT SwitchIO.xLiftCylinderRetractButton THEN
			SwitchIO.xLiftCylinderExtend:=1;
			SwitchIO.xLiftCylinderRetract:=0;
		END_IF;
		IF NOT SwitchIO.xLiftCylinderExtendButton AND  SwitchIO.xLiftCylinderRetractButton THEN
			SwitchIO.xLiftCylinderExtend:=0;
			SwitchIO.xLiftCylinderRetract:=1;
		END_IF;		
	END_IF;
END_FUNCTION_BLOCK
